   Button "Button_2" at 191,433 size 320x84; TextOff 'Testshot is active'
      Visibility <- "DB1900_IF_Robots_State_Robots{0}_TestShotRunning"
   Button "Template_Button_41" at 16,724 size 68x66; TextOff 'Text'; PictureList "Ico_navigation_2"; PictureOff "Setting_Nav_7"; Authorization "User administration"
      on Click: ActivateScreen("0035_Robot Setting", 0)
      ProcessValue <- "Nav_7"
      Visibility <- "NavUserChange"

screen "0035_Robot Setting" 1280x800, template "Navigation"
   on GenerateScreen: SetBit("DB1900_IF_Robots_Read"); SetBit("DB1901_Config_Robots_Read")
   Button "b_Incress_Pump_Setting" at 789,105 size 46x32; TextOff 'Text'; PictureOff "right arrow"
      on Click: function_dd21b452("DB613_Komponent_State_ReadDeviceNo", 1); function_dd21b452("DB612_Tank_State.ReadDeviceNo", 1)
   Button "b_Decress_Pump_Setting" at 269,105 size 46x32; TextOff 'Text'; PictureOff "left arrow"
      on Click: function_b9b71300("DB613_Komponent_State_ReadDeviceNo", 1); function_b9b71300("DB612_Tank_State.ReadDeviceNo", 1)
   Button "Button_2" at 124,176 size 480x580; TextOff 'Text'
   TextField "Text field_1" at 170,214 size 60x22; Text 'Robot:'
   TextField "Text field_2" at 170,251 size 50x22; Text 'KUKA'
   TextField "Text field_3" at 170,294 size 42x22; Text 'ABB'
   TextField "Text field_4" at 170,337 size 54x22; Text 'Fanuc'
   TextField "Text field_5" at 170,382 size 80x22; Text 'Motoman'
   TextField "Text field_6" at 168,428 size 149x22; Text 'Safety controller'
   TextField "Text field_7" at 170,472 size 107x22; Text 'Sync Switch'
   TextField "Text field_8" at 170,518 size 85x22; Text 'Shotware'
   TextField "Text field_9" at 170,564 size 78x22; Text 'Tracking'
   TextField "Text field_10" at 170,610 size 77x22; Text 'Testshot'
   TextField "Text field_11" at 170,656 size 77x22; Text 'Testshot'
   Button "Button_3" at 652,500 size 480x256; TextOff 'Text'
      Visibility <- "Robot Screen Visibility Control"
   TextField "Text field_12" at 682,531 size 179x22; Text 'Mixinghead Cleaning'
      Visibility <- "Robot Screen Visibility Control"
   TextField "Text field_13" at 678,573 size 42x22; Text 'LFI'
      Visibility <- "Robot Screen Visibility Control"
   TextField "Text field_14" at 678,616 size 90x22; Text 'Wet Clean'
      Visibility <- "Robot Screen Visibility Control"
   TextField "Text field_15" at 678,659 size 91x22; Text 'IR Station'
      Visibility <- "Robot Screen Visibility Control"
   TextField "Text field_16" at 678,702 size 54x22; Text 'Spare'
      Visibility <- "Robot Screen Visibility Control"
   TextField "Text field_17" at 930,573 size 106x22; Text 'Spray Clean'
      Visibility <- "Robot Screen Visibility Control"
   TextField "Text field_18" at 930,616 size 117x22; Text 'Brush station'
      Visibility <- "Robot Screen Visibility Control"
   TextField "Text field_19" at 930,659 size 108x22; Text 'Air Cleaning'
      Visibility <- "Robot Screen Visibility Control"
   TextField "Text field_20" at 930,702 size 54x22; Text 'Spare'
      Visibility <- "Robot Screen Visibility Control"
   Button "Check_Pump_WithFeedingPump" at 800,569 size 45x30; TextOff 'Text'; PictureOff "download"; PictureList "Check_Uncheck"
      on Click: InvertBit("DB1901_Config_Robots_Config_Robots{0}_With_Wet_Cleaning_LFI")
      Visibility <- "Robot Screen Visibility Control"
      ProcessValue <- "DB1901_Config_Robots_Config_Robots{0}_With_Wet_Cleaning_LFI"
   Button "Check_Pump_WithFeedingPump_1" at 800,612 size 45x30; TextOff 'Text'; PictureOff "download"; PictureList "Check_Uncheck"
      on Click: InvertBit("DB1901_Config_Robots_Config_Robots{0}_With_Wet_Cleaning")
      Visibility <- "Robot Screen Visibility Control"
      ProcessValue <- "DB1901_Config_Robots_Config_Robots{0}_With_Wet_Cleaning"
   Button "Check_Pump_WithFeedingPump_2" at 800,655 size 45x30; TextOff 'Text'; PictureOff "download"; PictureList "Check_Uncheck"
      on Click: InvertBit("DB1901_Config_Robots_Config_Robots{0}_With_IR_Station")
      Visibility <- "Robot Screen Visibility Control"
      ProcessValue <- "DB1901_Config_Robots_Config_Robots{0}_With_IR_Station"
   Button "Check_Pump_WithFeedingPump_3" at 800,698 size 45x30; TextOff 'Text'; PictureOff "download"; PictureList "Check_Uncheck"
      on Click: InvertBit("DB1901_Config_Robots_Config_Robots{0}_With_Belt_Filter")
      Visibility <- "Robot Screen Visibility Control"
      ProcessValue <- "DB1901_Config_Robots_Config_Robots{0}_With_Belt_Filter"
   Button "Check_Pump_WithFeedingPump_4" at 1057,569 size 45x30; TextOff 'Text'; PictureOff "download"; PictureList "Check_Uncheck"
      on Click: InvertBit("DB1901_Config_Robots_Config_Robots{0}_With_Wet_Cleaning_Spray")
      Visibility <- "Robot Screen Visibility Control"
      ProcessValue <- "DB1901_Config_Robots_Config_Robots{0}_With_Wet_Cleaning_Spray"
   Button "Check_Pump_WithFeedingPump_5" at 1057,612 size 45x30; TextOff 'Text'; PictureOff "download"; PictureList "Check_Uncheck"
      on Click: InvertBit("DB1901_Config_Robots_Config_Robots{0}_With_Brush_Station")
      Visibility <- "Robot Screen Visibility Control"
      ProcessValue <- "DB1901_Config_Robots_Config_Robots{0}_With_Brush_Station"
   Button "Check_Pump_WithFeedingPump_6" at 1057,655 size 45x30; TextOff 'Text'; PictureOff "download"; PictureList "Check_Uncheck"
      on Click: InvertBit("DB1901_Config_Robots_Config_Robots{0}_With_Air_Cleaner")
      Visibility <- "Robot Screen Visibility Control"
      ProcessValue <- "DB1901_Config_Robots_Config_Robots{0}_With_Air_Cleaner"
   Button "Check_Pump_WithFeedingPump_7" at 1057,698 size 45x30; TextOff 'Text'; PictureOff "download"; PictureList "Check_Uncheck"
      on Click: InvertBit("DB1901_Config_Robots_Config_Robots{0}_Spare_2_7")
      Visibility <- "Robot Screen Visibility Control"
      ProcessValue <- "DB1901_Config_Robots_Config_Robots{0}_Spare_2_7"
   Button "Check_Pump_WithFeedingPump_8" at 455,247 size 45x30; TextOff 'Text'; PictureOff "download"; PictureList "Check_Uncheck"
      on Click: InvertBit("DB1901_Config_Robots_Config_Robots{0}_Type_Kuka")
      ProcessValue <- "DB1901_Config_Robots_Config_Robots{0}_Type_Kuka"
   Button "Check_Pump_WithFeedingPump_9" at 455,290 size 45x30; TextOff 'Text'; PictureOff "download"; PictureList "Check_Uncheck"
      on Click: InvertBit("DB1901_Config_Robots_Config_Robots{0}_Type_ABB")
      ProcessValue <- "DB1901_Config_Robots_Config_Robots{0}_Type_ABB"
   Button "Check_Pump_WithFeedingPump_10" at 455,333 size 45x30; TextOff 'Text'; PictureOff "download"; PictureList "Check_Uncheck"
      on Click: InvertBit("DB1901_Config_Robots_Config_Robots{0}_Type_Fanuc")
      ProcessValue <- "DB1901_Config_Robots_Config_Robots{0}_Type_Fanuc"
   Button "Check_Pump_WithFeedingPump_11" at 455,378 size 45x30; TextOff 'Text'; PictureOff "download"; PictureList "Check_Uncheck"
      on Click: InvertBit("DB1901_Config_Robots_Config_Robots{0}_Type_Motoman")
      ProcessValue <- "DB1901_Config_Robots_Config_Robots{0}_Type_Motoman"
   Button "Check_Pump_WithFeedingPump_12" at 455,424 size 45x30; TextOff 'Text'; PictureOff "download"; PictureList "Check_Uncheck"
      on Click: InvertBit("DB1901_Config_Robots_Config_Robots{0}_With_Belt_Filter")
      ProcessValue <- "DB1901_Config_Robots_Config_Robots{0}_With_Belt_Filter"
   Button "Check_Pump_WithFeedingPump_13" at 455,468 size 45x30; TextOff 'Text'; PictureOff "download"; PictureList "Check_Uncheck"
      on Click: InvertBit("DB1901_Config_Robots_Config_Robots{0}_With_Synchronisation")
      ProcessValue <- "DB1901_Config_Robots_Config_Robots{0}_With_Synchronisation"
   Button "Check_Pump_WithFeedingPump_14" at 455,514 size 45x30; TextOff 'Text'; PictureOff "download"; PictureList "Check_Uncheck"
      on Click: InvertBit("DB1901_Config_Robots_Config_Robots{0}_With_Shotware")
      ProcessValue <- "DB1901_Config_Robots_Config_Robots{0}_With_Shotware"
   Button "Check_Pump_WithFeedingPump_15" at 455,560 size 45x30; TextOff 'Text'; PictureOff "download"; PictureList "Check_Uncheck"
      on Click: InvertBit("DB1901_Config_Robots_Config_Robots{0}_With_Tracking")
      ProcessValue <- "DB1901_Config_Robots_Config_Robots{0}_With_Tracking"
   Button "Check_Pump_WithFeedingPump_16" at 455,606 size 45x30; TextOff 'Text'; PictureOff "download"; PictureList "Check_Uncheck"
      on Click: InvertBit("DB1901_Config_Robots_Config_Robots{0}_With_Testshot")
      ProcessValue <- "DB1901_Config_Robots_Config_Robots{0}_With_Testshot"
   Button "Check_Pump_WithFeedingPump_17" at 455,652 size 45x30; TextOff 'Text'; PictureOff "download"; PictureList "Check_Uncheck"
      on Click: InvertBit("DB1901_Config_Robots_Config_Robots{0}_With_Cleaning")
      ProcessValue <- "DB1901_Config_Robots_Config_Robots{0}_With_Cleaning"
   Button "b_Pump_CoolingHeating" at 378,652 size 45x30; TextOff 'Text'; PictureOff "obeng"
      on Click: SetTag("Robot Screen Visibility Control", 1)
      Visibility <- "DB1901_Config_Robots_Config_Robots{0}_With_Cleaning"
   SymbolicIOField "Symbolic I/O field_1" at 326,104 size 451x32; TextOn '1'; TextOff '0'; TextList "Robot_name"
      ProcessValue <- "DB1900_IF_Robots_ReadWriteDeviceNo"
   Button "b_Close_Pump_CH" at 1080,502 size 51x41; TextOff 'Text'; PictureOff "images (1)"
      on Press: SetTag("Robot Screen Visibility Control", 0)
      Visibility <- "Robot Screen Visibility Control"

PopupScreen "Fault" 350x130
   on GenerateScreen: SetBit("PopUp_Restrict")
   Button "Button_1" at 262,89 size 53x32; TextOff 'Close'; PictureOff "images (7)"
      on Click: ResetBit("DB_MouldEditor_HMI_uData_sStatusBits_xFaultValuesnotvalid"); function_efd93a16("Fault", 446, 387, 0, -1, 1); ResetBit("PopUp_Restrict")
   Button "Button_2" at 186,88 size 53x32; TextOff 'Y'; PictureOff "_green_check.svg"
      on Click: ResetBit("DB_MouldEditor_HMI_uData_sStatusBits_xFaultValuesnotvalid"); ResetBit("DB_MouldEditor_HMI_uData_sStatusBits_xValueChanged"); function_efd93a16("Fault", 446, 387, 0, -1, 1); SetBit("DB_MouldEditor_HMI_uData_sStatusBits_xDiscardChanges"); ResetBit("PopUp_Restrict")
   TextField "Text field_1" at 96,37 size 145x40; Text 'Data Not Valid Unable to store !'
   GraphicView "Graphic view_1" at 19,36 size 47x40; Picture "Alarm Icon 1"

screen "Tes" 1280x800
   AlarmView "Alarm view_1" at 23,18 size 713x300
   Button "Button_1" at 23,350 size 119x63; TextOff 'Tes'
      on Press: "Custom_Datalog"()
   IOField "I/O field_1" at 426,450 size 96x32; FormatPattern 9999999999999999999999999999999999999999
      ProcessValue <- "tes_Time_1"
   IOField "I/O field_2" at 611,450 size 96x32; FormatPattern 9999999999999999999999999999999999999999
      ProcessValue <- "tes_Time_2"
   Button "Button_2" at 522,600 size 96x32; TextOff 'Tes Time'
      on Click: "Tes"()
   IOField "I/O field_3" at 522,536 size 96x32; FormatPattern 9999999999999999999999999999999999999999
      ProcessValue <- "tes_Time_3"
   IOField "I/O field_4" at 523,381 size 96x32; FormatPattern 9999999999999999999999999999999999999999
      ProcessValue <- "TP-Bereichszeiger_Date_Time_ActTime"
   TextField "Text field_1" at 542,351 size 58x22; Text 'Actual'
   TextField "Text field_2" at 527,510 size 87x22; Text 'Next time'
   TextField "Text field_3" at 444,423 size 61x22; Text 'Time 1'
   TextField "Text field_4" at 629,423 size 61x22; Text 'Time 2'
   DateTimeField "Date/time field_1" at 681,382 size 121x31
   AlarmView "Alarm view_2" at 34,635 size 809x165

screen "9020_Service" 1280x800, template "Navigation"
   on GenerateScreen: SetTag("ServiceScreenControl", 9020)
   Button "Button_3" at 326,104 size 451x32; TextOff 'Service'
   TextField "Text field_1" at 543,326 size 110x29; Text 'Contact :'
   TextField "Text field_2" at 413,374 size 370x29; Text 'Hotline: +49 (0) 89 - 8899 3152'
   TextField "Text field_3" at 434,423 size 329x29; Text 'Fax: +49 (0) 89 - 8899 4024'
   TextField "Text field_4" at 379,472 size 439x29; Text 'Email: serviceRPM@kraussmaffei.com'
   Button "MixingHeadButton_6" at 219,696 size 60x60; TextOff 'PLC IO MONITOR'; PictureList "ico_plcio"
      on Click: ActivateScreen("9021_Plc IO Monitor", 0)
      Appearance <- "ServiceScreenControl"
      ProcessValue <- "ServiceScreenControl"
   Button "MixingHeadButton_2" at 308,696 size 60x60; TextOff 'PLC IO MONITOR Web'; PictureOff "ico"; PictureList "ico_Web"
      on Click: ActivateScreen("9022_Web Explorer", 0)
      ProcessValue <- "ServiceScreenControl"
      Appearance <- "ServiceScreenControl"
   Button "MixingHeadButton_3" at 397,696 size 60x60; TextOff 'PLC IO MONITOR smart'; PictureList "ico_Smart"
      on Click: ActivateScreen("9023_SmartClient", 0)
      Appearance <- "ServiceScreenControl"
      ProcessValue <- "ServiceScreenControl"
   Button "MixingHeadButton_4" at 131,696 size 60x60; TextOff 'PLC IO MONITOR Service & Solutions'
      on Click: ActivateScreen("9020_Service", 0)
      Appearance <- "ServiceScreenControl"
   Button "MixingHeadButton_5" at 397,696 size 60x60; TextOff 'PLC IO MONITOR smart'
      on Click: ActivateScreen("9023_SmartClient", 0)
      Appearance <- "ServiceScreenControl"
      ProcessValue <- "ServiceScreenControl"
   Button "MixingHeadButton_7" at 308,696 size 60x60; TextOff 'PLC IO MONITOR Web'
      on Click: ActivateScreen("9022_Web Explorer", 0)
      ProcessValue <- "ServiceScreenControl"
      Appearance <- "ServiceScreenControl"
   Button "MixingHeadButton_8" at 219,696 size 60x60; TextOff 'PLC IO MONITOR'
      on Click: ActivateScreen("9021_Plc IO Monitor", 0)
      Appearance <- "ServiceScreenControl"
      ProcessValue <- "ServiceScreenControl"
   Button "MixingHeadButton_9" at 1060,696 size 60x60; TextOff 'DIAGNOSTIC'; PictureOff "information"; PictureList "ico_information"
      on Click: ActivateScreen("9029_Information", 0)
      Appearance <- "ServiceScreenControl"
      ProcessValue <- "ServiceScreenControl"
   Button "MixingHeadButton_1" at 486,696 size 60x60; TextOff 'DIAGNOSTIC'; PictureOff "Graphic_29"
      on Click: ActivateScreen("9024_Diagnostic Overview", 0); function_ce3c6af1("9024_Diagnostic Overview", "System diagnostics view_1")
      Appearance <- "ServiceScreenControl"

screen "9024_Diagnostic Overview" 1280x800, template "Navigation"
   on GenerateScreen: SetTag("ServiceScreenControl", 9024)
   Button "Button_3" at 326,104 size 451x32; TextOff 'Plc Variabel / Service'
   SysDiagControl "System diagnostics view_1" at 122,164 size 1032x518; InfoArea_RootNodeText 'Plant / Anlage'; BusyText 'Please Wait... / Bitte warten... / Please wait..........'; NavigationPath_RootText 'Diagnostic overview / Diagnose Überblick / Diagnostic Overview'
   Button "MixingHeadButton_6" at 219,696 size 60x60; TextOff 'PLC IO MONITOR'; PictureList "ico_plcio"
      on Click: ActivateScreen("9021_Plc IO Monitor", 0)
      Appearance <- "ServiceScreenControl"
      ProcessValue <- "ServiceScreenControl"
   Button "MixingHeadButton_1" at 486,696 size 60x60; TextOff 'DIAGNOSTIC'; PictureOff "Graphic_29"
      on Click: ActivateScreen("9024_Diagnostic Overview", 0); function_ce3c6af1("9024_Diagnostic Overview", "System diagnostics view_1")
      Appearance <- "ServiceScreenControl"
   Button "MixingHeadButton_2" at 308,696 size 60x60; TextOff 'PLC IO MONITOR Web'; PictureOff "ico"; PictureList "ico_Web"
      on Click: ActivateScreen("9022_Web Explorer", 0)
      ProcessValue <- "ServiceScreenControl"
      Appearance <- "ServiceScreenControl"
   Button "MixingHeadButton_3" at 397,696 size 60x60; TextOff 'PLC IO MONITOR smart'; PictureList "ico_Smart"
      on Click: ActivateScreen("9023_SmartClient", 0)
      Appearance <- "ServiceScreenControl"
      ProcessValue <- "ServiceScreenControl"
   Button "MixingHeadButton_5" at 397,696 size 60x60; TextOff 'PLC IO MONITOR smart'
      on Click: ActivateScreen("9023_SmartClient", 0)
      Appearance <- "ServiceScreenControl"
      ProcessValue <- "ServiceScreenControl"
   Button "MixingHeadButton_7" at 308,696 size 60x60; TextOff 'PLC IO MONITOR Web'
      on Click: ActivateScreen("9022_Web Explorer", 0)
      ProcessValue <- "ServiceScreenControl"
      Appearance <- "ServiceScreenControl"
   Button "MixingHeadButton_8" at 219,696 size 60x60; TextOff 'PLC IO MONITOR'
      on Click: ActivateScreen("9021_Plc IO Monitor", 0)
      Appearance <- "ServiceScreenControl"
      ProcessValue <- "ServiceScreenControl"
   Button "MixingHeadButton_9" at 1060,696 size 60x60; TextOff 'DIAGNOSTIC'; PictureOff "information"; PictureList "ico_information"
      on Click: ActivateScreen("9029_Information", 0)
      Appearance <- "ServiceScreenControl"
      ProcessValue <- "ServiceScreenControl"
   Button "MixingHeadButton_4" at 131,696 size 60x60; TextOff 'PLC IO MONITOR Service & Solutions'
      on Click: ActivateScreen("9020_Service", 0)
      Appearance <- "ServiceScreenControl"

screen "9022_Web Explorer" 1280x800, template "Navigation"
   on GenerateScreen: SetTag("ServiceScreenControl", 9022)
   HTMLBrowser "HTML browser_1" at 129,170 size 1021x509
   Button "Button_3" at 326,104 size 451x32; TextOff 'Plc Variabel / Service'
   Button "MixingHeadButton_6" at 219,696 size 60x60; TextOff 'PLC IO MONITOR'; PictureList "ico_plcio"
      on Click: ActivateScreen("9021_Plc IO Monitor", 0)
      Appearance <- "ServiceScreenControl"
      ProcessValue <- "ServiceScreenControl"
   Button "MixingHeadButton_2" at 308,696 size 60x60; TextOff 'PLC IO MONITOR Web'; PictureOff "ico"; PictureList "ico_Web"
      on Click: ActivateScreen("9022_Web Explorer", 0)
      ProcessValue <- "ServiceScreenControl"
      Appearance <- "ServiceScreenControl"
   Button "MixingHeadButton_3" at 397,696 size 60x60; TextOff 'PLC IO MONITOR smart'; PictureList "ico_Smart"
      on Click: ActivateScreen("9023_SmartClient", 0)
      Appearance <- "ServiceScreenControl"
      ProcessValue <- "ServiceScreenControl"
   Button "MixingHeadButton_5" at 397,696 size 60x60; TextOff 'PLC IO MONITOR smart'
      on Click: ActivateScreen("9023_SmartClient", 0)
      Appearance <- "ServiceScreenControl"
      ProcessValue <- "ServiceScreenControl"
   Button "MixingHeadButton_7" at 308,696 size 60x60; TextOff 'PLC IO MONITOR Web'
      on Click: ActivateScreen("9022_Web Explorer", 0)
      ProcessValue <- "ServiceScreenControl"
      Appearance <- "ServiceScreenControl"
   Button "MixingHeadButton_8" at 219,696 size 60x60; TextOff 'PLC IO MONITOR'
      on Click: ActivateScreen("9021_Plc IO Monitor", 0)
      Appearance <- "ServiceScreenControl"
      ProcessValue <- "ServiceScreenControl"
   Button "MixingHeadButton_9" at 1060,696 size 60x60; TextOff 'DIAGNOSTIC'; PictureOff "information"; PictureList "ico_information"
      on Click: ActivateScreen("9029_Information", 0)
      Appearance <- "ServiceScreenControl"
      ProcessValue <- "ServiceScreenControl"
   Button "MixingHeadButton_4" at 131,696 size 60x60; TextOff 'PLC IO MONITOR Service & Solutions'
      on Click: ActivateScreen("9020_Service", 0)
      Appearance <- "ServiceScreenControl"
   Button "MixingHeadButton_1" at 486,696 size 60x60; TextOff 'DIAGNOSTIC'; PictureOff "Graphic_29"
      on Click: ActivateScreen("9024_Diagnostic Overview", 0); function_ce3c6af1("9024_Diagnostic Overview", "System diagnostics view_1")
      Appearance <- "ServiceScreenControl"

screen "9023_SmartClient" 1280x800, template "Navigation"
   on GenerateScreen: SetTag("ServiceScreenControl", 9023)
   SmartClientView "Sm@rtClient view_1" at 121,111 size 1035x534
   Button "MixingHeadButton_6" at 219,696 size 60x60; TextOff 'PLC IO MONITOR'; PictureList "ico_plcio"
      on Click: ActivateScreen("9021_Plc IO Monitor", 0)
      Appearance <- "ServiceScreenControl"
      ProcessValue <- "ServiceScreenControl"
   Button "MixingHeadButton_2" at 308,696 size 60x60; TextOff 'PLC IO MONITOR Web'; PictureOff "ico"; PictureList "ico_Web"
      on Click: ActivateScreen("9022_Web Explorer", 0)
      ProcessValue <- "ServiceScreenControl"
      Appearance <- "ServiceScreenControl"
   Button "MixingHeadButton_3" at 397,696 size 60x60; TextOff 'PLC IO MONITOR smart'; PictureList "ico_Smart"
      on Click: ActivateScreen("9023_SmartClient", 0)
      Appearance <- "ServiceScreenControl"
      ProcessValue <- "ServiceScreenControl"
   Button "MixingHeadButton_5" at 397,696 size 60x60; TextOff 'PLC IO MONITOR smart'
      on Click: ActivateScreen("9023_SmartClient", 0)
      Appearance <- "ServiceScreenControl"
      ProcessValue <- "ServiceScreenControl"
   Button "MixingHeadButton_7" at 308,696 size 60x60; TextOff 'PLC IO MONITOR Web'
      on Click: ActivateScreen("9022_Web Explorer", 0)
      ProcessValue <- "ServiceScreenControl"
      Appearance <- "ServiceScreenControl"
   Button "MixingHeadButton_8" at 219,696 size 60x60; TextOff 'PLC IO MONITOR'
      on Click: ActivateScreen("9021_Plc IO Monitor", 0)
      Appearance <- "ServiceScreenControl"
      ProcessValue <- "ServiceScreenControl"
   Button "MixingHeadButton_9" at 1060,696 size 60x60; TextOff 'DIAGNOSTIC'; PictureOff "information"; PictureList "ico_information"
      on Click: ActivateScreen("9029_Information", 0)
      Appearance <- "ServiceScreenControl"
      ProcessValue <- "ServiceScreenControl"
   Button "MixingHeadButton_4" at 131,696 size 60x60; TextOff 'PLC IO MONITOR Service & Solutions'
      on Click: ActivateScreen("9020_Service", 0)
      Appearance <- "ServiceScreenControl"
   Button "MixingHeadButton_1" at 486,696 size 60x60; TextOff 'DIAGNOSTIC'; PictureOff "Graphic_29"
      on Click: ActivateScreen("9024_Diagnostic Overview", 0); function_ce3c6af1("9024_Diagnostic Overview", "System diagnostics view_1")
      Appearance <- "ServiceScreenControl"

screen "9029_Information" 1280x800, template "Navigation"
   on GenerateScreen: SetTag("ServiceScreenControl", 9029)
   Button "Button_3" at 326,104 size 451x32; TextOff 'Service'
   TextField "Text field_1" at 356,210 size 90x22; Text 'Customer:'
   TextField "Text field_2" at 356,248 size 127x22; Text 'Order number:'
   TextField "Text field_3" at 356,286 size 75x22; Text 'Version:'
   TextField "Text field_4" at 356,324 size 145x22; Text 'Production year:'
   TextField "Text field_5" at 356,362 size 147x22; Text 'Machine number:'
   TextField "Text field_6" at 356,400 size 207x22; Text 'Wiring diagram number:'
   TextField "Text field_7" at 356,438 size 135x22; Text 'Additional info:'
   TextField "Text field_8" at 356,476 size 135x22; Text 'Additional info:'
   TextField "Text field_9" at 356,514 size 135x22; Text 'Additional info:'
   TextField "Text field_10" at 356,552 size 135x22; Text 'Additional info:'
   TextField "Text field_11" at 356,590 size 135x22; Text 'Additional info:'
   IOField "I/O field_1" at 563,200 size 351x32; FormatPattern ?????????????????????????????????????????????
      ProcessValue <- "Customer"
      Visibility <- "NavUserChange"
   IOField "I/O field_2" at 564,238 size 146x32; FormatPattern ?????????????????????????????????????????????
      ProcessValue <- "Order_number"
      Visibility <- "NavUserChange"
   IOField "I/O field_3" at 565,276 size 86x32; FormatPattern ?????????????????????????????????????????????
      ProcessValue <- "Version"
      Visibility <- "NavUserChange"
   IOField "I/O field_4" at 566,314 size 105x32; FormatPattern ?????????????????????????????????????????????
      ProcessValue <- "Production_year"
      Visibility <- "NavUserChange"
   IOField "I/O field_5" at 567,352 size 156x32; FormatPattern ?????????????????????????????????????????????
      ProcessValue <- "Machine_number"
      Visibility <- "NavUserChange"
   IOField "I/O field_6" at 568,390 size 155x32; FormatPattern ?????????????????????????????????????????????
      ProcessValue <- "Wiring_diagram_number"
      Visibility <- "NavUserChange"
   IOField "I/O field_7" at 569,428 size 351x32; FormatPattern ?????????????????????????????????????????????
      ProcessValue <- "Additional_info_1"
      Visibility <- "NavUserChange"
   IOField "I/O field_8" at 570,466 size 351x32; FormatPattern ?????????????????????????????????????????????
      ProcessValue <- "Additional_info_2"
      Visibility <- "NavUserChange"
   IOField "I/O field_9" at 571,504 size 351x32; FormatPattern ?????????????????????????????????????????????
      ProcessValue <- "Additional_info_3"
      Visibility <- "NavUserChange"
   IOField "I/O field_10" at 572,542 size 351x32; FormatPattern ?????????????????????????????????????????????
      ProcessValue <- "Additional_info_4"
      Visibility <- "NavUserChange"
   IOField "I/O field_11" at 573,580 size 351x32; FormatPattern ?????????????????????????????????????????????
      ProcessValue <- "Additional_info_5"
      Visibility <- "NavUserChange"
   Button "MixingHeadButton_6" at 219,696 size 60x60; TextOff 'PLC IO MONITOR'; PictureList "ico_plcio"
      on Click: ActivateScreen("9021_Plc IO Monitor", 0)
      Appearance <- "ServiceScreenControl"
      ProcessValue <- "ServiceScreenControl"
   Button "MixingHeadButton_2" at 308,696 size 60x60; TextOff 'PLC IO MONITOR Web'; PictureOff "ico"; PictureList "ico_Web"
      on Click: ActivateScreen("9022_Web Explorer", 0)
      ProcessValue <- "ServiceScreenControl"
      Appearance <- "ServiceScreenControl"
   Button "MixingHeadButton_3" at 397,696 size 60x60; TextOff 'PLC IO MONITOR smart'; PictureList "ico_Smart"
      on Click: ActivateScreen("9023_SmartClient", 0)
      Appearance <- "ServiceScreenControl"
      ProcessValue <- "ServiceScreenControl"
   Button "MixingHeadButton_5" at 397,696 size 60x60; TextOff 'PLC IO MONITOR smart'
      on Click: ActivateScreen("9023_SmartClient", 0)
      Appearance <- "ServiceScreenControl"
      ProcessValue <- "ServiceScreenControl"
   Button "MixingHeadButton_7" at 308,696 size 60x60; TextOff 'PLC IO MONITOR Web'
      on Click: ActivateScreen("9022_Web Explorer", 0)
      ProcessValue <- "ServiceScreenControl"
      Appearance <- "ServiceScreenControl"
   Button "MixingHeadButton_8" at 219,696 size 60x60; TextOff 'PLC IO MONITOR'
      on Click: ActivateScreen("9021_Plc IO Monitor", 0)
      Appearance <- "ServiceScreenControl"
      ProcessValue <- "ServiceScreenControl"
   Button "MixingHeadButton_9" at 1060,696 size 60x60; TextOff 'DIAGNOSTIC'; PictureOff "information"; PictureList "ico_information"
      on Click: ActivateScreen("9029_Information", 0)
      Appearance <- "ServiceScreenControl"
      ProcessValue <- "ServiceScreenControl"
   Button "MixingHeadButton_10" at 1058,400 size 60x60; TextOff 'DIAGNOSTIC From SD'; PictureOff "information"; PictureList "ico_information"
      ProcessValue <- "ServiceScreenControl"
      Visibility <- "NavUserChange"
   Button "MixingHeadButton_11" at 1056,578 size 60x60; TextOff 'DIAGNOSTIC From USB'; PictureOff "information"; PictureList "ico_information"
      ProcessValue <- "ServiceScreenControl"
   Button "MixingHeadButton_4" at 131,696 size 60x60; TextOff 'PLC IO MONITOR Service & Solutions'
      on Click: ActivateScreen("9020_Service", 0)
      Appearance <- "ServiceScreenControl"
   Button "MixingHeadButton_1" at 486,696 size 60x60; TextOff 'DIAGNOSTIC'; PictureOff "Graphic_29"
      on Click: ActivateScreen("9024_Diagnostic Overview", 0); function_ce3c6af1("9024_Diagnostic Overview", "System diagnostics view_1")
      Appearance <- "ServiceScreenControl"

screen "0038_RFID" 1280x800, template "Navigation"
   TextField "Text field_1" at 564,156 size 112x22; Text 'RFID Reader'
   TextField "Text field_2" at 274,202 size 47x22; Text 'MH 1'
   TextField "Text field_3" at 870,202 size 47x22; Text 'MH 2'

VB script "ScreenOpen"
   'Tip:
   ' 1. Use the <CTRL+SPACE> or <CTRL+I> shortcut to open a list of all objects and functions
   ' 2. Write the code using the HMI Runtime object.
   '  Example: HmiRuntime.Screens("Screen_1").
   ' 3. Use the <CTRL+J> shortcut to create an object reference.
   'Write the code as of this position:
   
   
   
   
   
   Select Case SmartTags("Navigation_7")
   	Case 1
   		'Open Screen Machine Setting
   		bec8f1e5-2ab1-45f6-ad91-1d37c469eb91 1000_General Machine Configuration,1000
   		b21d3eaf-4e31-425c-ad1a-ba4e4002cacc Navigation_7,0
   		
   	Case 2
   		'Open Screen Pump Setting
   		bec8f1e5-2ab1-45f6-ad91-1d37c469eb91 0012_Pump Setting,12
   		b21d3eaf-4e31-425c-ad1a-ba4e4002cacc Navigation_7,0
   	Case 3
   		'Open Screen Tank Setting
   		bec8f1e5-2ab1-45f6-ad91-1d37c469eb91 0007_Tank Setting,7
   		b21d3eaf-4e31-425c-ad1a-ba4e4002cacc Navigation_7,0
   	Case 4
   		'open screen MH Setting
   		bec8f1e5-2ab1-45f6-ad91-1d37c469eb91 0005_Mixinghead Settting,3
   		b21d3eaf-4e31-425c-ad1a-ba4e4002cacc Navigation_7,0
   		
   	Case 5
   		'Open Mixinghead hydraulic setting
   		b21d3eaf-4e31-425c-ad1a-ba4e4002cacc MixingHead Options,1
   		b21d3eaf-4e31-425c-ad1a-ba4e4002cacc Navigation_7,0
   		
   	Case 6 
   		'Open Robot Setting
   		bec8f1e5-2ab1-45f6-ad91-1d37c469eb91 0035_Robot Setting,35
   		b21d3eaf-4e31-425c-ad1a-ba4e4002cacc Navigation_7,0
   	Case Else
   		'statementblock_n
   End Select
   
   
   	

VB script "ToolAllocation_First"
   Select Case SmartTags("DB939_Tool_alloc_HMI_AllocList_page")
   Case 2
   		b21d3eaf-4e31-425c-ad1a-ba4e4002cacc Tool_Allocation_Numb_1,31
   		b21d3eaf-4e31-425c-ad1a-ba4e4002cacc Tool_Allocation_Numb_2,32
   		b21d3eaf-4e31-425c-ad1a-ba4e4002cacc Tool_Allocation_Numb_3,33
   		b21d3eaf-4e31-425c-ad1a-ba4e4002cacc Tool_Allocation_Numb_4,34
   		b21d3eaf-4e31-425c-ad1a-ba4e4002cacc Tool_Allocation_Numb_5,35
   		b21d3eaf-4e31-425c-ad1a-ba4e4002cacc Tool_Allocation_Numb_6,36
   		b21d3eaf-4e31-425c-ad1a-ba4e4002cacc Tool_Allocation_Numb_7,37
   		b21d3eaf-4e31-425c-ad1a-ba4e4002cacc Tool_Allocation_Numb_8,38
   		b21d3eaf-4e31-425c-ad1a-ba4e4002cacc Tool_Allocation_Numb_9,39
   		b21d3eaf-4e31-425c-ad1a-ba4e4002cacc Tool_Allocation_Numb_10,40
   		b21d3eaf-4e31-425c-ad1a-ba4e4002cacc Tool_Allocation_Numb_11,41
   		b21d3eaf-4e31-425c-ad1a-ba4e4002cacc Tool_Allocation_Numb_12,42
   		b21d3eaf-4e31-425c-ad1a-ba4e4002cacc Tool_Allocation_Numb_13,43
   		b21d3eaf-4e31-425c-ad1a-ba4e4002cacc Tool_Allocation_Numb_14,44
   		b21d3eaf-4e31-425c-ad1a-ba4e4002cacc Tool_Allocation_Numb_15,45
   		
   		'KANAN
   		b21d3eaf-4e31-425c-ad1a-ba4e4002cacc Tool_Allocation_Numb_16,46
   		b21d3eaf-4e31-425c-ad1a-ba4e4002cacc Tool_Allocation_Numb_17,47
   		b21d3eaf-4e31-425c-ad1a-ba4e4002cacc Tool_Allocation_Numb_18,48
   		b21d3eaf-4e31-425c-ad1a-ba4e4002cacc Tool_Allocation_Numb_19,49
   		b21d3eaf-4e31-425c-ad1a-ba4e4002cacc Tool_Allocation_Numb_20,50
   		b21d3eaf-4e31-425c-ad1a-ba4e4002cacc Tool_Allocation_Numb_21,51
   		b21d3eaf-4e31-425c-ad1a-ba4e4002cacc Tool_Allocation_Numb_22,52
   		b21d3eaf-4e31-425c-ad1a-ba4e4002cacc Tool_Allocation_Numb_23,53
   		b21d3eaf-4e31-425c-ad1a-ba4e4002cacc Tool_Allocation_Numb_24,54
   		b21d3eaf-4e31-425c-ad1a-ba4e4002cacc Tool_Allocation_Numb_25,55
   		b21d3eaf-4e31-425c-ad1a-ba4e4002cacc Tool_Allocation_Numb_26,56
   		b21d3eaf-4e31-425c-ad1a-ba4e4002cacc Tool_Allocation_Numb_27,57
   		b21d3eaf-4e31-425c-ad1a-ba4e4002cacc Tool_Allocation_Numb_28,58
   		b21d3eaf-4e31-425c-ad1a-ba4e4002cacc Tool_Allocation_Numb_29,59
   		b21d3eaf-4e31-425c-ad1a-ba4e4002cacc Tool_Allocation_Numb_30,60		
   Case 3
   		b21d3eaf-4e31-425c-ad1a-ba4e4002cacc Tool_Allocation_Numb_1,61
   		b21d3eaf-4e31-425c-ad1a-ba4e4002cacc Tool_Allocation_Numb_2,62
   		b21d3eaf-4e31-425c-ad1a-ba4e4002cacc Tool_Allocation_Numb_3,63
   		b21d3eaf-4e31-425c-ad1a-ba4e4002cacc Tool_Allocation_Numb_4,64
   		b21d3eaf-4e31-425c-ad1a-ba4e4002cacc Tool_Allocation_Numb_5,65
   		b21d3eaf-4e31-425c-ad1a-ba4e4002cacc Tool_Allocation_Numb_6,66
   		b21d3eaf-4e31-425c-ad1a-ba4e4002cacc Tool_Allocation_Numb_7,67
   		b21d3eaf-4e31-425c-ad1a-ba4e4002cacc Tool_Allocation_Numb_8,68
   		b21d3eaf-4e31-425c-ad1a-ba4e4002cacc Tool_Allocation_Numb_9,69
   		b21d3eaf-4e31-425c-ad1a-ba4e4002cacc Tool_Allocation_Numb_10,70
   		b21d3eaf-4e31-425c-ad1a-ba4e4002cacc Tool_Allocation_Numb_11,71
   		b21d3eaf-4e31-425c-ad1a-ba4e4002cacc Tool_Allocation_Numb_12,72
   		b21d3eaf-4e31-425c-ad1a-ba4e4002cacc Tool_Allocation_Numb_13,73
   		b21d3eaf-4e31-425c-ad1a-ba4e4002cacc Tool_Allocation_Numb_14,74
   		b21d3eaf-4e31-425c-ad1a-ba4e4002cacc Tool_Allocation_Numb_15,75